// TIA Portal project "DHARMA_1500" (V15)

(* hardware
DEVICE "HMI_DHARMA"  TP1200 Comfort
   slot 0: "KraussMaffeiHMI"  TP1200 Comfort  6AV2 124-0MC01-0AX0  14.0.1.0
   slot 1: "HMI_RT_1"  TP1200 Comfort  6AV2 124-0MC01-0AX0  14.0.1.0
   slot 5: "KraussMaffeiHMI.IE_CP_1"  PROFINET Interface  14.0.1.0
      slot 1: "PROFINET Interface_1"  PROFINET Interface
         slot 1: "Port_1"  Port
         slot 2: "Port_2"  Port
   slot 7: "KraussMaffeiHMI.MPI/DP_CP_1"  MPI/DP Interface  14.0.1.0
DEVICE "S71500/ET200MP station_1"  S7-1500 station
   slot 0: "Rail_0"  Rack  6ES7 590-1***0-0AA0
   slot 1: "PLC_DHARMA"  CPU 1515-2 PN  6ES7 515-2AM01-0AB0  V2.5
      slot 3: "CPU display_1"  6ES7591-1BA00-0AA0
*)

// ===== PLC "PLC_DHARMA"  CPU 1515-2 PN =====

VAR_GLOBAL   // PLC tag table "Standard-Variablentabelle"
   "Sensor_CupIsAtTestshotposition" AT %I18.7 : Bool;   // The cup is at the testhotposition
   "PAW_800_tool_1" AT %QW800 : Word;
   "Tag_3" AT %Q13.2 : Bool;
   "Tag_4" AT %Q13.3 : Bool;
   "Duese_K2_MH01" AT %Q51.2 : Bool;
   "HF_pulse_alarm_GWK1" AT %M1002.4 : Bool;
   "FP_temperingunit_off" AT %M1002.5 : Bool;
   "FP_temperingunit_on" AT %M1002.6 : Bool;
   "With_MC03" AT %M710.0 : Bool;
   "With_MC04" AT %M710.1 : Bool;
   "HF_pulse_alarm_GWK2" AT %M1002.7 : Bool;
   "HF_new_setvalue_Of_ShotData" AT %M701.2 : Bool;
   "HM_Shotend" AT %M50.0 : Bool;
   "TIM_FRA_WDG3" AT %T15 : Timer;
   "TIM_FRA_WDG4" AT %T16 : Timer;
   "T_CupIsAtTestshotposition" AT %T192 : Timer;
END_VAR

VAR_GLOBAL CONSTANT   // PLC tag table "Standard-Variablentabelle"
   "AmountPartShots" : Int := 8;   // Array lenght for UDT 925
   "AmountToolsDB" : Int := 100;   // Array lenght for each DB
   "AmountAllocationAutomatic" : Int := 210;   // Array lenght for DB931 (always 30 Steps)
   "AmountTools" : Int := 200;   // Array lenght for DB930
END_VAR

VAR_GLOBAL   // PLC tag table "E/A- Belegung INput"
   "F_Klima" AT %I4.7 : Bool;   // Malfunction air-condition
   "P_Vacuum_C1" AT %I117.0 : Bool;   // Vacuum reached componet 1
   "P_Vacuum_C2" AT %I117.1 : Bool;   // Vacuum reached componet 2
   "S_BarrelDetection_C1" AT %I111.0 : Bool;   // Special: Barrel exist for the component 1
   "S_BarrelDetection_C2" AT %I112.0 : Bool;   // Special: Barrel exist for the component 2
   "F_Fan_Pump_C1" AT %I110.0 : Bool;   // Fault fuse fan pump component 1
   "F_Fan_Pump_C2" AT %I110.1 : Bool;   // Fault fuse fan pump component 2
   "F_FCFeedingP_C1" AT %I110.4 : Bool;   // Fault frequency drive feed pump component 1
   "F_FCFeedingP_C2" AT %I110.5 : Bool;   // Fault frequency drive feed pump component 2
   "T_Start_Test_C1" AT %I26.3 : Bool;   // Start button for test component 1
   "T_Start_Test_C2" AT %I27.3 : Bool;   // Start button for test component 1
   "T_Stop_Test" AT %I27.2 : Bool;   // Stop button for test component
   "S_OM_Test" AT %I26.2 : Bool;   // Switch for selection operation mode test
   "P_2_MK_Hydr" AT %I2.5 : Bool;   // hydraulic pressure 2 reached
   "ES_GBE_C1" AT %I1.7 : Bool;   // Emergency stop from nucleation component 1
   "F_GBE_C1" AT %I0.5 : Bool;   // Fault Supply nucleation component 1
   "F_GBE_Faulty_C1" AT %I0.6 : Bool;   // Fault Message from nuvleation component 1
   "F_GBE_Ready_C1" AT %I1.3 : Bool;   // Nucleation ready component 1
   "F_FeedPump_C2" AT %I8.6 : Bool;   // Fault filling pump daytank component 2
   "S_DryRun_Feed_C1" AT %I119.2 : Bool;   // Dry run protection feeding pump tank component 1
   "S_DryRun_Feed_C2" AT %I118.3 : Bool;   // Dry run protection feeding pump tank component 2
   "Container_FaultSupply" AT %I10.7 : Bool;   // Faulty power supply containerstaion
   "ES_Door_Robot_01" AT %I13.2 : Bool;   // Emergency stop door robot 1
   "ES_Door_TestShot_01" AT %I18.4 : Bool;   // Emergency stop door testshot robot 1
   "ES_Container_C1" AT %I10.5 : Bool;   // Emergency stop from containerstaion component 1
   "TestShot_MouldExist" AT %I14.4 : Bool;   // Testshot: Mould existing
   "TestShot_Level" AT %I14.5 : Bool;   // Testshot: Filling level
   "S_SelectDoor_Robot_01" AT %I13.0 : Bool;   // Select open door robot 1
   "AS_Door_Robot_01" AT %I13.3 : Bool;   // Automatic stop door robot 1
   "S_QuittDoor_Robot_01" AT %I13.1 : Bool;   // Quitt automatic stop door robot 1
   "S_SelectDoor_TestShot_01" AT %I18.0 : Bool;   // Select open door test shot 1
   "AS_Door_TestShot_01" AT %I18.3 : Bool;   // Automatic stop door test shot 1
   "S_QuittDoor_TestShot_01" AT %I18.1 : Bool;   // Quitt automatic stop door test shot 1
   "AS_RobotInArea1" AT %I12.0 : Bool;   // Save Move (EPS) area 1
   "AS_RobotInArea2" AT %I12.1 : Bool;   // Save Move (EPS) area 2
   "AS_Dryside" AT %I8.7 : Bool;   // Automatic stop from mould carrier 01
   "AS" AT %I12.7 : Bool;   // Emergency stop from dryside
   "F_CoolingDevice" AT %I0.4 : Bool;   // Faulty supply chiller
   "Container_Ready_C1" AT %I10.1 : Bool;   // Signal container is ready for filling daytank component 1
   "Container_Ready_C2" AT %I10.2 : Bool;   // Signal container is ready for filling daytank component 2
   "Container_Fillpump_run_C1" AT %I10.3 : Bool;   // Signal container filling pump is running component 1
   "Container_Fillpump_run_C2" AT %I10.4 : Bool;   // Signal container filling pump is running component 2
   "Container_Faulty" AT %I10.6 : Bool;   // Signal container fault existing
   "F_TraceHeatingM1_C3" AT %I17.3 : Bool;
   "F_FeedingP_C1" AT %I24.0 : Bool;   // Fault Feeding pump component 1
   "F_FeedingP_C2" AT %I25.0 : Bool;   // Fault Feeding pump component 2
   "F_SupplyHeatingM1" AT %I16.0 : Bool;   // Stoerung versorgung heizung
   "F_TraceHeatingM1_C1" AT %I16.1 : Bool;   // Stoerung begleitheizung vorlauf ruecklauf poly
   "F_TraceHeatingM1_C2" AT %I16.2 : Bool;   // Stoerung begleitheizung vorlauf ruecklauf iso
   "F_TraceHeatingM1_C1_2" AT %I16.3 : Bool;
   "F_TraceHeatingM1_C2_2" AT %I16.4 : Bool;
   "F_Robot_01" AT %I12.6 : Bool;   // Fault fuse robot 01
   "F_Airdryer" AT %I0.1 : Bool;   // Fault Airdryer
   "ES_Extern(SGM_or_MC)" AT %I0.0 : Bool;   // Emergency stop from extern (SGM or Mould carrier)
   "F_Fuse_Machine" AT %I0.2 : Bool;   // Fault circuit breakes machine component 1/2
   "F_Fuse_MH" AT %I0.3 : Bool;   // Fault fuse mixinghead
   "ES_Operatingpanel" AT %I1.5 : Bool;   // Emergency stop control panel PUC 08
   "ES_Machine" AT %I1.4 : Bool;   // Emergency stop machine component 1/2
   "Controlvoltage" AT %I0.7 : Bool;   // Control voltage on
   "ES_Robot_01" AT %I12.5 : Bool;   // Emergency stop from robot 01
   "ES_Central" AT %I1.6 : Bool;   // Emergency stop from central
   "S_OM_Manual" AT %I1.0 : Bool;   // Operating mode manual
   "S_OM_Auto" AT %I1.1 : Bool;   // Operating mode automatic
   "T_QuitFault" AT %I1.2 : Bool;
   "F_MK_Hydr" AT %I2.0 : Bool;   // malfunction hydraulicmotor
   "F_Fil_MK_Hydr_VL" AT %I2.1 : Bool;   // hydraulic filter polluted forwardslauf
   "L_Min_Oel_MK_Hydr" AT %I2.2 : Bool;   // hydraulic fill level OK
   "C_Max_Oel_MK_Hydr" AT %I2.3 : Bool;   // Max temperature hydraulic
   "P_MK_Hydr" AT %I2.4 : Bool;   // hydraulic pressure reached
   "C_Cooling_Hydr" AT %I2.6 : Bool;   // Start cooling hydraulic
   "F_Heating" AT %I2.7 : Bool;   // Fault Heating Day tank
   "Select_door_TT" AT %I120.5 : Bool;
   "AS_door_TT" AT %I120.3 : Bool;
   "Quit_door_TT" AT %I120.4 : Bool;
   "F_fuse_vacuum_pump_Seg_1" AT %I121.4 : Bool;
   "F_fuse_vacuum_pump_Seg_2" AT %I122.4 : Bool;
   "F_fuse_vacuum_pump_Seg_3" AT %I123.4 : Bool;
   "F_fuse_vacuum_pump_Seg_4" AT %I124.4 : Bool;
   "Safety_switch_MC_1" AT %I121.2 : Bool;
   "Safety_switch_MC_2" AT %I122.2 : Bool;
   "Safety_switch_MC_3" AT %I123.2 : Bool;
   "Safety_switch_MC_4" AT %I124.2 : Bool;
   "S_Start_TestShot_01" AT %I18.2 : Bool;   // Start automatic test shot 1
   "AS_RobotInArea3" AT %I12.2 : Bool;   // Save Move (EPS) area 3
   "AS_RobotInArea4" AT %I12.3 : Bool;   // Save Move (EPS) area 4
   "AS_RobotInArea5" AT %I18.5 : Bool;   // Save Move (EPS) area 5
   "AS_RobotInArea6" AT %I18.6 : Bool;   // Save Move (EPS) area 6
   "AS_Lightbarrier_back_MC01" AT %I30.3 : Bool;   // Automatic stop light barrier behind MC 1
   "ES_MC02" AT %I30.4 : Bool;   // Emergency stop from mould carrier 2
   "AS_tool_exists_MC02" AT %I30.5 : Bool;   // Automatic stop tool exists mould carrier 2
   "AS_MC02" AT %I30.6 : Bool;   // Automatic stop from mould carrier 2
   "AS_Lightbarrier_back_MC02" AT %I30.7 : Bool;   // Automatic stop light barrier behind MC 2
   "ES_MC03" AT %I31.0 : Bool;   // Emergency stop from mould carrier 3
   "AS_tool_exists_MC03" AT %I31.1 : Bool;   // Automatic stop tool exists mould carrier 3
   "AS_MC03" AT %I31.2 : Bool;   // Automatic stop from mould carrier 3
   "AS_Lightbarrier_back_MC03" AT %I31.3 : Bool;   // Automatic stop light barrier behind MC 3
   "ES_MC04" AT %I31.4 : Bool;   // Emergency stop from mould carrier 4
   "AS_tool_exists_MC04" AT %I31.5 : Bool;   // Automatic stop tool exists mould carrier 4
   "AS_MC04" AT %I31.6 : Bool;   // Automatic stop from mould carrier 4
   "AS_Lightbarrier_back_MC04" AT %I31.7 : Bool;   // Automatic stop light barrier behind MC 4
   "ES_MC01" AT %I30.0 : Bool;   // Emergency stop from mould carrier 1
   "AS_tool_exists_MC01" AT %I30.1 : Bool;   // Automatic stop tool exists mould carrier 1
   "AS_MC01" AT %I30.2 : Bool;   // Automatic stop from mould carrier 1
   "P_air" AT %I19.7 : Bool;   // Pressure air inlet
   "C_Start_Refill_POLY_ON" AT %Q11.1 : Bool;
   "C_Start_Refill_ISO_ON" AT %Q11.2 : Bool;
   "Release_door_TT" AT %Q120.1 : Bool;
   "Selected_door_TT" AT %Q120.0 : Bool;
   "O_vacuum_pump_Seg_1" AT %Q121.1 : Bool;
   "O_vacuum_pump_Seg_2" AT %Q121.2 : Bool;
   "O_vacuum_pump_Seg_3" AT %Q121.3 : Bool;
   "O_vacuum_pump_Seg_4" AT %Q121.4 : Bool;
   "FHM_Takt_Verz_RT1" AT %M900.0 : Bool;
   "HM_FP_Takt_Verz_RT1" AT %M900.1 : Bool;
END_VAR

VAR_GLOBAL   // PLC tag table "E/A- Belegung OUTput"
   "K_ControllVoltageOff" AT %Q0.4 : Bool;
   "K_Stoerung_FT" AT %Q3.0 : Bool;   // malfunction to mouldcarrier
   "K_Schussende_FT" AT %Q3.1 : Bool;   // Shotend an mouldcarrier
   "H_CP_Back_MH1" AT %Q3.2 : Bool;   // MH01: indicator cleaning piston back
   "H_Rel_Foaming_MH1" AT %Q3.3 : Bool;   // MH01: indicator release foaming
   "H_HighPressure_MH1" AT %Q3.4 : Bool;   // MH01: indicator high pressure circulation
   "V_MH_open_MH1" AT %Q115.0 : Bool;   // MH00: Valve mixinghead open
   "V_CP_Forward_MH1" AT %Q115.1 : Bool;   // MH00: valve cleaning piston forward
   "V_PumpVacuum_C1" AT %Q117.0 : Bool;
   "V_PressureVacuum_C1" AT %Q117.1 : Bool;
   "V_PumpVacuum_C2" AT %Q117.2 : Bool;
   "V_PressureVacuum_C2" AT %Q117.3 : Bool;
   "M_CirculationPump_C3" AT %Q118.0 : Bool;   // Circulation Pump net component 3
   "V_PumpVacuum_C3" AT %Q117.4 : Bool;
   "V_PressureVacuum_C3" AT %Q117.5 : Bool;
   "V_PressureVacuum_C4" AT %Q117.7 : Bool;
   "V_Inert_MH1" AT %Q122.6 : Bool;   // MH01: Valve Nitrogen for Inerting
   "V_Inert_Piston_MH1" AT %Q131.5 : Bool;   // MH01: Valve Nitrogen Piston
   "M_Fan_Pump_Net_C1" AT %Q110.0 : Bool;   // Fan pump net component 1
   "M_Fan_Pump_Net_C2" AT %Q110.1 : Bool;   // Fan pump net component 2
   "M_FeedingP_Start_C1" AT %Q24.1 : Bool;   // Feedingpump release frequency drive component 1
   "M_FeedingP_Start_C2" AT %Q25.1 : Bool;   // Feedingpump release frequency drive component 2
   "V_Test_C1" AT %Q26.2 : Bool;   // Valve for test component 1
   "V_Test_C2" AT %Q27.2 : Bool;   // Valve for test component 2
   "H_Test_C1" AT %Q26.3 : Bool;   // Visual information for test component 1
   "H_Test_C2" AT %Q27.3 : Bool;   // Visual information for test component 2
   "V_Pump_2Point_C1" AT %Q5.0 : Bool;   // 2 Point adjustment component pump component 1
   "M_FeedPump_C1" AT %Q27.0 : Bool;   // Valve for feedpump Daytank Component 1
   "M_FeedPump_C2" AT %Q26.0 : Bool;   // Valve for feedpump Daytank Component 2
   "V_Pump_2Point_C2" AT %Q5.1 : Bool;   // 2 Point adjustment component pump component 2
   "V_OpenDoor_Robot_01" AT %Q13.1 : Bool;   // Clamping valve door robot 01
   "H_ReleaseDoor_Robot_01" AT %Q13.0 : Bool;   // Light door robot 01
   "V_OpenDoor_TestShot_01" AT %Q18.0 : Bool;   // Clamping valve door test shot 01
   "H_AutoStopQuit" AT %Q0.3 : Bool;   // Indicator auto stop acknowledged
   "H_ReleaseDoor_TestShot_01" AT %Q18.1 : Bool;   // Light door test shot 01
   "V_P_builtup_MH_Hydr_M1" AT %Q1.1 : Bool;   // Hydraulic pressur built up mixinhead 1
   "V_Cooling_Hydr" AT %Q1.2 : Bool;   // Hydraulic 1 valve for oil cooling
   "M_MH_Hydr_Net_M1" AT %Q1.0 : Bool;   // Hydraulic motor net mixinghead 1
   "H_Fault_lamp_M1" AT %Q0.0 : Bool;   // Visual fault warning M1
   "H_Fault_horn_M1" AT %Q0.1 : Bool;   // Acustical fault warning M1
   "H_Ready_for_Operation" AT %Q0.2 : Bool;
   "H_TestShot_active_01" AT %Q18.2 : Bool;   // Automatic test shot is running 01
END_VAR

VAR_GLOBAL   // PLC tag table "I/O- Pentan"
   "E_Voralarm_Pentan" AT %I116.0 : Bool;   // Pentan: Pre alarm (20%) pentan
   "P_Voralarm_Stickstoff" AT %I116.1 : Bool;   // Pentan: Pre alarm nitrogen
   "P_Alarm_Stickstoff" AT %I116.2 : Bool;   // Pentan: Alarm nitrogen
   "P_Alarm_VersorgungN" AT %I116.3 : Bool;   // Pentan: Alarm nitrogen supply
   "E_Absaugung_bereit" AT %I116.4 : Bool;   // Pentan: Exhaust system ready
   "E_Pentanpumpe_laeuft" AT %I116.5 : Bool;   // Pentan: Pump pentan running
   "E_Pentamix_Ready" AT %I116.6 : Bool;   // Pentan: Pentamix ready for supply
   "ES_Pentamix" AT %I116.7 : Bool;
   "P_Nitrogen_Inerting_OK" AT %I17.6 : Bool;   // Nitrogen pressure for Inerting ok
   "Flow_Nitrogen Inert_OK" AT %I17.7 : Bool;   // Nitrogen flow after start inerting ok
   "K_Machine_Running" AT %Q116.0 : Bool;   // Pentan: Signal machine running to gas warning desk
   "K_Request_WeekendMode" AT %Q116.1 : Bool;   // Pentan: Request for weekend mode to gas warning desk
   "V_Fass_Pentan1" AT %Q1101.6 : Bool;
   "V_ChargingTank_C1_2" AT %Q22.4 : Bool;   // Filling valve 2 tank component 1
END_VAR

VAR_GLOBAL   // PLC tag table "I/O- PN Modul Flow Output"
   "V_ChargingTank_C2_2" AT %Q22.3 : Bool;   // Filling valve 2 tank component 1
   "M_Pump_Net_C1" AT %Q20.0 : Bool;   // Pump net componet 1
   "M_Pump_Start_C1" AT %Q20.1 : Bool;   // Pump release frequency drive component 1
   "M_Platefilter_C1" AT %Q20.7 : Bool;   // Platefilter net componet 1
   "M_Pump_Net_C2" AT %Q22.0 : Bool;   // Pump net component 2
   "M_Pump_Start_C2" AT %Q22.1 : Bool;   // Pump release frequency drive component 2
   "M_Platefilter_C2" AT %Q22.7 : Bool;   // Platefilter net component 2
   "V_HP_Heater_Cooling_C1" AT %Q21.6 : Bool;   // Valve for cooling high pressure heatexchanger component 1
   "V_HP_Heater_Bypass_C1" AT %Q80.6 : Bool;   // Valve for bypass high pressure heatexchanger component 1
   "V_HP_Heater_Cooling_C2" AT %Q23.6 : Bool;   // Valve for cooling high pressure heatexchanger component 2
   "K_Filling_Tank_C2_TL" AT %Q23.7 : Bool;   // Potential-free contact for filling Tank component 2 from another source
   "M_FU_Start_RW_K1" AT %Q21.1 : Bool;   // Agitator release frequency drive component 1
   "M_FU_Start_RW_K2" AT %Q23.1 : Bool;   // Agitator release frequency drive component 2
   "M_FeedingP_C1" AT %Q24.0 : Bool;   // Feeding pump net component 2
   "M_FeedingP_C2" AT %Q25.0 : Bool;   // Feeding pump net component 2
   "K_Filling_Tank_C2" AT %Q23.3 : Bool;   // Potential-free contact for filling Tank component 2
   "K_Filling_Tank_C1" AT %Q21.3 : Bool;   // Potential-free contact for filling Tank component 1
   "M_AgitatorBarrel_C1" AT %Q20.4 : Bool;   // Agitator barrel net component 1
   "M_Agitator_C1" AT %Q21.0 : Bool;   // Agitator net component 1
   "K_HeatingTank_C1" AT %Q20.2 : Bool;   // Heating Day tank net componet 1
   "V_Coolingwater_C1" AT %Q21.4 : Bool;   // Valve cooling water tank component 1
   "V_ChargingTank_C1" AT %Q21.2 : Bool;   // Filling valve tank component 1
   "V_Barrel_C1" AT %Q20.5 : Bool;   // Valve barrel station component 1
   "V_Heatexchanger_C1" AT %Q21.5 : Bool;   // heat exchangerValve Poly
   "V_Barrel_C2" AT %Q22.5 : Bool;   // Valve barrel station component 2
   "V_Heatexchanger_C2" AT %Q23.5 : Bool;   // heat exchangerValve component 2
   "V_Coolingwater_C2" AT %Q23.4 : Bool;   // Valve cooling water component 2
   "K_HeatingTank_C2" AT %Q22.2 : Bool;   // Heating Day tank net componet 2
   "V_ChargingTank_C2" AT %Q23.2 : Bool;   // Filling valve component 2
   "M_Agitator_C2" AT %Q23.0 : Bool;   // Agitator net component 2
   "V_LowPressure_Circ_C1" AT %Q20.6 : Bool;   // Low pressure circulation component 1
   "V_LowPressure_Circ_C2" AT %Q22.6 : Bool;   // Low pressure circulation component 2
END_VAR

VAR_GLOBAL   // PLC tag table "I/O- PN Modul Flow Input"
   "F_FC_Pump_C1" AT %I20.2 : Bool;   // Fault frequency drive componet 1
   "F_Pump_C1" AT %I20.3 : Bool;   // Fault pump componet 1
   "P_Prepressure_Pump_C1" AT %I20.4 : Bool;   // Pre pressure pump componet 1
   "P_Min_C1" AT %I20.5 : Bool;   // Min. pressure pump componet 1
   "P_Max_C1" AT %I20.6 : Bool;   // Max. pressure pump componet 1
   "F_Platefilter_C1" AT %I20.7 : Bool;   // Fault Platefilter component 1
   "F_FC_Agitator_C1" AT %I21.1 : Bool;   // Malfunction frequency converter agitator component 1
   "F_FC_Pump_C2" AT %I22.2 : Bool;   // Fault frequency drive componet 2
   "F_Pump_C2" AT %I22.3 : Bool;   // Fault pump componet 2
   "P_Prepressure_Pump_C2" AT %I22.4 : Bool;   // Pre pressure pump componet 2
   "P_Min_C2" AT %I22.5 : Bool;   // Min. pressure pump componet 2
   "F_Platefilter_C2" AT %I22.7 : Bool;   // Fault Platefilter component 2
   "P_Max_C2" AT %I22.6 : Bool;   // Max. pressure pump componet 2
   "F_FC_Agitator_C2" AT %I23.1 : Bool;   // Malfunction frequency converter agitator component 2
   "F_Agitator_C1" AT %I21.0 : Bool;   // Fault agitator componet 1
   "F_Temperiergeraet_C1" AT %I21.7 : Bool;   // Malfunction temperature stabilizer component 1
   "L_Tank_min_C1" AT %I21.2 : Bool;   // Min fill level tank componet 1
   "L_Tank_start_C1" AT %I21.3 : Bool;   // Start refilling level tank componet 1
   "L_Tank_stop_C1" AT %I21.4 : Bool;   // Stop refilling level tank componet 1
   "L_DT_max_C1" AT %I21.5 : Bool;   // Max. Filling level componet 1
   "L_DripTray_C1" AT %I21.6 : Bool;   // Max. level drip tray componet 1
   "F_Agitator_C2" AT %I23.0 : Bool;   // Fault agitator componet 2
   "F_Temperiergeraet_C2" AT %I23.7 : Bool;   // Malfunction temperature stabilizer component 2
   "L_Tank_min_C2" AT %I23.2 : Bool;   // Min fill level componet 2
   "L_Tank_start_C2" AT %I23.3 : Bool;   // Start refilling level componet 2
   "L_Tank_stop_C2" AT %I23.4 : Bool;   // Stop refilling level componet 2
   "L_DT_max_C2" AT %I23.5 : Bool;   // Max. Filling level componet 2
   "L_DripTray_C2" AT %I23.6 : Bool;   // Max. level drip tray componet 2
   "Kracht_C1_A_Flowrate" AT %I20.0 : Bool;
   "Kracht_C1_B_Flowrate" AT %I20.1 : Bool;
   "Kracht_C2_A_Flowrate" AT %I22.0 : Bool;
   "Kracht_C2_B_Flowrate" AT %I22.1 : Bool;
END_VAR

VAR_GLOBAL   // PLC tag table "I/O- PN Modul Mixinghead Output"
   "V_SWU_MH01" AT %Q50.5 : Bool;   // MH01: Valve switch over unit
   "H_Shotcounter_MH01" AT %Q52.7 : Bool;   // MH01: shot counter
   "V_CP_Forward_MH01" AT %Q50.4 : Bool;   // MH01: valve cleaning piston forward
   "H_CP_Back_MH01" AT %Q52.4 : Bool;   // MH01: indicator cleaning piston back
   "H_Rel_Foaming_MH01" AT %Q52.6 : Bool;   // MH01: indicator release foaming
   "H_HighPressure_MH01" AT %Q52.5 : Bool;   // MH01: indicator high pressure circulation
   "K_Fault_MC01" AT %Q50.6 : Bool;   // MH01: malfunction PU-machine to mouldcarrier
   "K_ShotEnd_MC01" AT %Q50.7 : Bool;   // MH01: Shotend PU-machine to mouldcarrier
   "V_MH_open_MH01" AT %Q50.0 : Bool;   // MH01: Valve mixinghead open
   "V_LowPressure_Circ_MH01" AT %Q53.7 : Bool;   // MH01: low pressure circulation Poly/ Iso
   "V_MH_open_MH02" AT %Q54.0 : Bool;   // MH01: Valve mixinghead open
   "V_CP_Forward_MH02" AT %Q54.4 : Bool;   // MH01: valve cleaning piston forward
   "V_SWU_MH02" AT %Q54.5 : Bool;   // MH01: Valve switch over unit
   "K_Fault_MC02" AT %Q54.6 : Bool;   // MH01: malfunction PU-machine to mouldcarrier
   "K_ShotEnd_MC02" AT %Q54.7 : Bool;   // MH01: Shotend PU-machine to mouldcarrier
   "H_CP_Back_MH02" AT %Q56.4 : Bool;   // MH01: indicator cleaning piston back
   "H_HighPressure_MH02" AT %Q56.5 : Bool;   // MH01: indicator high pressure circulation
   "H_Rel_Foaming_MH02" AT %Q56.6 : Bool;   // MH01: indicator release foaming
   "H_Shotcounter_MH02" AT %Q56.7 : Bool;   // MH01: shot counter
   "V_LowPressure_Circ_MH02" AT %Q57.7 : Bool;   // MH01: low pressure circulation Poly/ Iso
   "V_MH_open_MH03" AT %Q58.0 : Bool;   // MH01: Valve mixinghead open
   "V_CP_Forward_MH03" AT %Q58.4 : Bool;   // MH01: valve cleaning piston forward
   "V_SWU_MH03" AT %Q58.5 : Bool;   // MH01: Valve switch over unit
   "K_Fault_MC03" AT %Q58.6 : Bool;   // MH01: malfunction PU-machine to mouldcarrier
   "K_ShotEnd_MC03" AT %Q58.7 : Bool;   // MH01: Shotend PU-machine to mouldcarrier
   "H_CP_Back_MH03" AT %Q60.4 : Bool;   // MH01: indicator cleaning piston back
   "H_HighPressure_MH03" AT %Q60.5 : Bool;   // MH01: indicator high pressure circulation
   "H_Rel_Foaming_MH03" AT %Q60.6 : Bool;   // MH01: indicator release foaming
   "H_Shotcounter_MH03" AT %Q60.7 : Bool;   // MH01: shot counter
   "V_LowPressure_Circ_MH03" AT %Q61.7 : Bool;   // MH01: low pressure circulation Poly/ Iso
   "V_MH_open_MH04" AT %Q62.0 : Bool;   // MH01: Valve mixinghead open
   "V_CP_Forward_MH04" AT %Q62.4 : Bool;   // MH01: valve cleaning piston forward
   "V_SWU_MH04" AT %Q62.5 : Bool;   // MH01: Valve switch over unit
   "K_Fault_MC04" AT %Q62.6 : Bool;   // MH01: malfunction PU-machine to mouldcarrier
   "K_ShotEnd_MC04" AT %Q62.7 : Bool;   // MH01: Shotend PU-machine to mouldcarrier
   "H_CP_Back_MH04" AT %Q64.4 : Bool;   // MH01: indicator cleaning piston back
   "H_HighPressure_MH04" AT %Q64.5 : Bool;   // MH01: indicator high pressure circulation
   "H_Rel_Foaming_MH04" AT %Q64.6 : Bool;   // MH01: indicator release foaming
   "H_Shotcounter_MH04" AT %Q64.7 : Bool;   // MH01: shot counter
   "V_LowPressure_Circ_MH04" AT %Q65.7 : Bool;   // MH01: low pressure circulation Poly/ Iso
   "V_MH_open_MH05" AT %Q66.0 : Bool;   // MH01: Valve mixinghead open
   "V_CP_Forward_MH05" AT %Q66.4 : Bool;   // MH01: valve cleaning piston forward
   "V_SWU_MH05" AT %Q66.5 : Bool;   // MH01: Valve switch over unit
   "K_Fault_MC05" AT %Q66.6 : Bool;   // MH01: malfunction PU-machine to mouldcarrier
   "K_ShotEnd_MC05" AT %Q66.7 : Bool;   // MH01: Shotend PU-machine to mouldcarrier
   "H_CP_Back_MH05" AT %Q68.4 : Bool;   // MH01: indicator cleaning piston back
   "H_HighPressure_MH05" AT %Q68.5 : Bool;   // MH01: indicator high pressure circulation
   "H_Rel_Foaming_MH05" AT %Q68.6 : Bool;   // MH01: indicator release foaming
   "H_Shotcounter_MH05" AT %Q68.7 : Bool;   // MH01: shot counter
   "V_LowPressure_Circ_MH05" AT %Q69.7 : Bool;   // MH01: low pressure circulation Poly/ Iso
   "V_MH_open_MH06" AT %Q70.0 : Bool;   // MH01: Valve mixinghead open
   "V_CP_Forward_MH06" AT %Q70.4 : Bool;   // MH01: valve cleaning piston forward
   "V_SWU_MH06" AT %Q70.5 : Bool;   // MH01: Valve switch over unit
   "K_Fault_MC06" AT %Q70.6 : Bool;   // MH01: malfunction PU-machine to mouldcarrier
   "K_ShotEnd_MC06" AT %Q70.7 : Bool;   // MH01: Shotend PU-machine to mouldcarrier
   "H_CP_Back_MH06" AT %Q72.4 : Bool;   // MH01: indicator cleaning piston back
   "H_HighPressure_MH06" AT %Q72.5 : Bool;   // MH01: indicator high pressure circulation
   "H_Rel_Foaming_MH06" AT %Q72.6 : Bool;   // MH01: indicator release foaming
   "H_Shotcounter_MH06" AT %Q72.7 : Bool;   // MH01: shot counter
   "V_LowPressure_Circ_MH06" AT %Q73.7 : Bool;   // MH01: low pressure circulation Poly/ Iso
   "V_MH_open_MH07" AT %Q74.0 : Bool;   // MH01: Valve mixinghead open
   "V_CP_Forward_MH07" AT %Q74.4 : Bool;   // MH01: valve cleaning piston forward
   "V_SWU_MH07" AT %Q74.5 : Bool;   // MH01: Valve switch over unit
   "K_Fault_MC07" AT %Q74.6 : Bool;   // MH01: malfunction PU-machine to mouldcarrier
   "K_ShotEnd_MC07" AT %Q74.7 : Bool;   // MH01: Shotend PU-machine to mouldcarrier
   "H_CP_Back_MH07" AT %Q76.4 : Bool;   // MH01: indicator cleaning piston back
   "H_HighPressure_MH07" AT %Q76.5 : Bool;   // MH01: indicator high pressure circulation
   "H_Rel_Foaming_MH07" AT %Q76.6 : Bool;   // MH01: indicator release foaming
   "H_Shotcounter_MH07" AT %Q76.7 : Bool;   // MH01: shot counter
   "V_LowPressure_Circ_MH07" AT %Q77.7 : Bool;   // MH01: low pressure circulation Poly/ Iso
   "V_MH_open_MH08" AT %Q78.0 : Bool;   // MH01: Valve mixinghead open
   "V_CP_Forward_MH08" AT %Q78.4 : Bool;   // MH01: valve cleaning piston forward
   "V_SWU_MH08" AT %Q78.5 : Bool;   // MH01: Valve switch over unit
   "K_Fault_MC08" AT %Q78.6 : Bool;   // MH01: malfunction PU-machine to mouldcarrier
   "K_ShotEnd_MC08" AT %Q78.7 : Bool;   // MH01: Shotend PU-machine to mouldcarrier
   "H_CP_Back_MH08" AT %Q80.4 : Bool;   // MH01: indicator cleaning piston back
   "H_HighPressure_MH08" AT %Q80.5 : Bool;   // MH01: indicator high pressure circulation
   "K_Filling_Tank_C1_TL" AT %Q21.7 : Bool;   // Potential-free contact for filling Tank component 1 from another source
   "H_Shotcounter_MH08" AT %Q80.7 : Bool;   // MH01: shot counter
   "V_LowPressure_Circ_MH08" AT %Q81.7 : Bool;   // MH01: low pressure circulation Poly/ Iso
   "V_MH_open_MH09" AT %Q82.0 : Bool;   // MH01: Valve mixinghead open
   "V_CP_Forward_MH09" AT %Q82.4 : Bool;   // MH01: valve cleaning piston forward
   "V_SWU_MH09" AT %Q82.5 : Bool;   // MH01: Valve switch over unit
   "K_Fault_MC09" AT %Q82.6 : Bool;   // MH01: malfunction PU-machine to mouldcarrier
   "K_ShotEnd_MC09" AT %Q82.7 : Bool;   // MH01: Shotend PU-machine to mouldcarrier
   "H_CP_Back_MH09" AT %Q84.4 : Bool;   // MH01: indicator cleaning piston back
   "H_HighPressure_MH09" AT %Q84.5 : Bool;   // MH01: indicator high pressure circulation
   "H_Rel_Foaming_MH09" AT %Q84.6 : Bool;   // MH01: indicator release foaming
   "H_Shotcounter_MH09" AT %Q84.7 : Bool;   // MH01: shot counter
   "V_LowPressure_Circ_MH09" AT %Q85.7 : Bool;   // MH01: low pressure circulation Poly/ Iso
   "V_MH_open_MH10" AT %Q86.0 : Bool;   // MH01: Valve mixinghead open
   "V_CP_Forward_MH10" AT %Q86.4 : Bool;   // MH01: valve cleaning piston forward
   "V_SWU_MH10" AT %Q86.5 : Bool;   // MH01: Valve switch over unit
   "K_Fault_MC10" AT %Q86.6 : Bool;   // MH01: malfunction PU-machine to mouldcarrier
   "K_ShotEnd_MC10" AT %Q86.7 : Bool;   // MH01: Shotend PU-machine to mouldcarrier
   "H_CP_Back_MH10" AT %Q88.4 : Bool;   // MH01: indicator cleaning piston back
   "H_HighPressure_MH10" AT %Q88.5 : Bool;   // MH01: indicator high pressure circulation
   "H_Rel_Foaming_MH10" AT %Q88.6 : Bool;   // MH01: indicator release foaming
   "H_Shotcounter_MH10" AT %Q88.7 : Bool;   // MH01: shot counter
   "V_LowPressure_Circ_MH10" AT %Q95.7 : Bool;   // MH01: low pressure circulation Poly/ Iso
   "V_Bypass_C1" AT %Q51.1 : Bool;
   "V_Bypass_C2" AT %Q51.3 : Bool;
   "Duese_K1_MH01" AT %Q51.0 : Bool;
END_VAR

VAR_GLOBAL   // PLC tag table "I/O- PN Modul Mixinghead Input"
   "T_CP_forward_MH01" AT %I52.3 : Bool;   // MH01: Button cleaning piston forwards
   "T_CP_back_MH01" AT %I52.4 : Bool;   // MH01: Button cleaning piston back
   "S_ProgrNo_Bit40_MH01" AT %I51.6 : Bool;   // MH01: preselection program no. *10 MH BIT 2
   "P_Min_Air" AT %I53.6 : Bool;   // MH01: Min. Druck Reinigungsluft
   "P_Max_Air" AT %I53.7 : Bool;   // MH01: Max. Druck Reinigungsluft
   "S_ProgrNo_Bit80_MH01" AT %I51.7 : Bool;   // MH01: preselection program no. *10 MH BIT 3
   "ES_OP_Panel_MH01" AT %I50.2 : Bool;   // MH01: Emergency stop operating panel mixinghead
   "IPS_MH_MH01" AT %I50.0 : Bool;   // MH01: Inductive proximity switch mixinghead
   "IPS_CP_MH01" AT %I50.1 : Bool;   // MH01: Inductive proximity switch cleaning piston mixinghead
   "K_PreparationFoamingMC01" AT %I50.6 : Bool;   // MH01: preparation foaming from mouldcarrier
   "K_FoamingReleaseMC01" AT %I50.7 : Bool;   // MH01: shot release from mouldcarrier
   "S_Rel_SWU_MH01" AT %I52.2 : Bool;   // MH01: release switch over unit
   "S_Manuel_MH01" AT %I52.0 : Bool;   // MH01: operation mode manual
   "S_Automatic_MH01" AT %I52.1 : Bool;   // MH01: operation mode automatic
   "T_Highpressure_MH01" AT %I52.5 : Bool;   // MH01: Button high pressure circulation
   "S_ProgrNo_Bit20_MH01" AT %I51.5 : Bool;   // MH01: preselection program no. *10 MH BIT 1
   "S_ProgrNo_Bit10_MH01" AT %I51.4 : Bool;   // MH01: preselection program no. *10 MH BIT 0
   "S_ProgNoSelectMH01" AT %IB51 : Byte;   // MH01: preselection program no. MH
   "S_ProgrNo_Bit0_MH01" AT %I51.0 : Bool;   // MH01: preselection program no. MH BIT 0
   "S_ProgrNo_Bit1_MH01" AT %I51.1 : Bool;   // MH01: preselection program no. MH BIT 1
   "S_ProgrNo_Bit2_MH01" AT %I51.2 : Bool;   // MH01: preselection program no. MH BIT 2
   "S_ProgrNo_Bit3_MH01" AT %I51.3 : Bool;   // MH01: preselection program no. MH BIT 3
   "T_Start_MH01" AT %I52.6 : Bool;   // MH01: Button Start foaming
   "T_Stop_MH01" AT %I52.7 : Bool;   // MH01: Button Stop foaming
   "T_BreakeOpen_MH01" AT %I53.5 : Bool;   // MH01: Button to open the boom brake
   "IPS_MH_MH02" AT %I54.0 : Bool;   // MH02: Inductive proximity switch mixinghead
   "IPS_CP_MH02" AT %I54.1 : Bool;   // MH02: Inductive proximity switch cleaning piston mixinghead
   "ES_OP_Panel_MH02" AT %I54.2 : Bool;   // MH02: Emergency stop operating panel mixinghead
   "K_PreparationFoamingMC02" AT %I54.6 : Bool;   // MH02: preparation foaming from mouldcarrier
   "K_FoamingReleaseMC02" AT %I54.7 : Bool;   // MH02: shot release from mouldcarrier
   "S_ProgNoSelectMH02" AT %IB55 : Byte;   // MH02: preselection program no. MH
   "S_ProgrNo_Bit0_MH02" AT %I55.0 : Bool;   // MH02: preselection program no. MH BIT 0
   "S_ProgrNo_Bit1_MH02" AT %I55.1 : Bool;   // MH02: preselection program no. MH BIT 1
   "S_ProgrNo_Bit2_MH02" AT %I55.2 : Bool;   // MH02: preselection program no. MH BIT 2
   "S_ProgrNo_Bit3_MH02" AT %I55.3 : Bool;   // MH02: preselection program no. MH BIT 3
   "S_ProgrNo_Bit10_MH02" AT %I55.4 : Bool;   // MH02: preselection program no. *10 MH BIT 0
   "S_ProgrNo_Bit20_MH02" AT %I55.5 : Bool;   // MH02: preselection program no. *10 MH BIT 1
   "S_ProgrNo_Bit40_MH02" AT %I55.6 : Bool;   // MH02: preselection program no. *10 MH BIT 2
   "S_ProgrNo_Bit80_MH02" AT %I55.7 : Bool;   // MH02: preselection program no. *10 MH BIT 3
   "S_Manuel_MH02" AT %I724.0 : Bool;   // MH02: operation mode manual
   "S_Automatic_MH02" AT %I724.1 : Bool;   // MH02: operation mode automatic
   "S_Rel_SWU_MH02" AT %I724.2 : Bool;   // MH02: release switch over unit
   "T_CP_forward_MH02" AT %I724.3 : Bool;   // MH02: Button cleaning piston forwards
   "T_CP_back_MH02" AT %I724.4 : Bool;   // MH02: Button cleaning piston back
   "T_Highpressure_MH02" AT %I724.5 : Bool;   // MH02: Button high pressure circulation
   "T_Start_MH02" AT %I724.6 : Bool;   // MH02: Button Start foaming
   "T_Stop_MH02" AT %I724.7 : Bool;   // MH02: Button Stop foaming
   "P_Min_Air_MH02" AT %I725.6 : Bool;   // MH02: Min. Druck Reinigungsluft
   "P_Max_Air_MH02" AT %I725.7 : Bool;   // MH02: Max. Druck Reinigungsluft
   "T_BreakeOpen_MH02" AT %I725.5 : Bool;   // MH02: Button to open the boom brake
   "IPS_MH_MH03" AT %I726.0 : Bool;   // MH03: Inductive proximity switch mixinghead
   "IPS_CP_MH03" AT %I726.1 : Bool;   // MH03: Inductive proximity switch cleaning piston mixinghead
   "ES_OP_Panel_MH03" AT %I726.2 : Bool;   // MH03: Emergency stop operating panel mixinghead
   "K_PreparationFoamingMC03" AT %I726.6 : Bool;   // MH03: preparation foaming from mouldcarrier
   "K_FoamingReleaseMC03" AT %I726.7 : Bool;   // MH03: shot release from mouldcarrier
   "S_ProgNoSelectMH03" AT %IB727 : Byte;   // MH03: preselection program no. MH
   "S_ProgrNo_Bit0_MH03" AT %I727.0 : Bool;   // MH03: preselection program no. MH BIT 0
   "S_ProgrNo_Bit1_MH03" AT %I727.1 : Bool;   // MH03: preselection program no. MH BIT 1
   "S_ProgrNo_Bit2_MH03" AT %I727.2 : Bool;   // MH03: preselection program no. MH BIT 2
   "S_ProgrNo_Bit3_MH03" AT %I727.3 : Bool;   // MH03: preselection program no. MH BIT 3
   "S_ProgrNo_Bit10_MH03" AT %I727.4 : Bool;   // MH03: preselection program no. *10 MH BIT 0
   "S_ProgrNo_Bit20_MH03" AT %I727.5 : Bool;   // MH03: preselection program no. *10 MH BIT 1
   "S_ProgrNo_Bit40_MH03" AT %I727.6 : Bool;   // MH03: preselection program no. *10 MH BIT 2
   "S_ProgrNo_Bit80_MH03" AT %I727.7 : Bool;   // MH03: preselection program no. *10 MH BIT 3
   "S_Manuel_MH03" AT %I728.0 : Bool;   // MH03: operation mode manual
   "S_Automatic_MH03" AT %I728.1 : Bool;   // MH03: operation mode automatic
   "S_Rel_SWU_MH03" AT %I728.2 : Bool;   // MH03: release switch over unit
   "T_CP_forward_MH03" AT %I728.3 : Bool;   // MH03: Button cleaning piston forwards
   "T_CP_back_MH03" AT %I728.4 : Bool;   // MH03: Button cleaning piston back
   "T_Highpressure_MH03" AT %I728.5 : Bool;   // MH03: Button high pressure circulation
   "T_Start_MH03" AT %I728.6 : Bool;   // MH03: Button Start foaming
   "T_Stop_MH03" AT %I728.7 : Bool;   // MH03: Button Stop foaming
   "P_Min_Air_MH03" AT %I729.6 : Bool;   // MH03: Min. Druck Reinigungsluft
   "P_Max_Air_MH03" AT %I729.7 : Bool;   // MH03: Max. Druck Reinigungsluft
   "T_BreakeOpen_MH03" AT %I729.5 : Bool;   // MH03: Button to open the boom brake
   "IPS_MH_MH04" AT %I730.0 : Bool;   // MH03: Inductive proximity switch mixinghead
   "IPS_CP_MH04" AT %I730.1 : Bool;   // MH03: Inductive proximity switch cleaning piston mixinghead
   "ES_OP_Panel_MH04" AT %I730.2 : Bool;   // MH03: Emergency stop operating panel mixinghead
   "K_PreparationFoamingMC04" AT %I730.6 : Bool;   // MH03: preparation foaming from mouldcarrier
   "K_FoamingReleaseMC04" AT %I730.7 : Bool;   // MH03: shot release from mouldcarrier
   "S_ProgNoSelectMH04" AT %IB731 : Byte;   // MH03: preselection program no. MH
   "S_ProgrNo_Bit0_MH04" AT %I731.0 : Bool;   // MH03: preselection program no. MH BIT 0
   "S_ProgrNo_Bit1_MH04" AT %I731.1 : Bool;   // MH03: preselection program no. MH BIT 1
   "S_ProgrNo_Bit2_MH04" AT %I731.2 : Bool;   // MH03: preselection program no. MH BIT 2
   "S_ProgrNo_Bit3_MH04" AT %I731.3 : Bool;   // MH03: preselection program no. MH BIT 3
   "S_ProgrNo_Bit10_MH04" AT %I731.4 : Bool;   // MH03: preselection program no. *10 MH BIT 0
   "S_ProgrNo_Bit20_MH04" AT %I731.5 : Bool;   // MH03: preselection program no. *10 MH BIT 1
   "S_ProgrNo_Bit40_MH04" AT %I731.6 : Bool;   // MH03: preselection program no. *10 MH BIT 2
   "S_ProgrNo_Bit80_MH04" AT %I731.7 : Bool;   // MH03: preselection program no. *10 MH BIT 3
   "S_Manuel_MH04" AT %I732.0 : Bool;   // MH03: operation mode manual
   "S_Automatic_MH04" AT %I732.1 : Bool;   // MH03: operation mode automatic
   "S_Rel_SWU_MH04" AT %I732.2 : Bool;   // MH03: release switch over unit
   "T_CP_forward_MH04" AT %I732.3 : Bool;   // MH03: Button cleaning piston forwards
   "T_CP_back_MH04" AT %I732.4 : Bool;   // MH03: Button cleaning piston back
   "T_Highpressure_MH04" AT %I732.5 : Bool;   // MH03: Button high pressure circulation
   "T_Start_MH04" AT %I732.6 : Bool;   // MH03: Button Start foaming
   "T_Stop_MH04" AT %I732.7 : Bool;   // MH03: Button Stop foaming
   "P_Min_Air_MH04" AT %I733.6 : Bool;   // MH03: Min. Druck Reinigungsluft
   "P_Max_Air_MH04" AT %I733.7 : Bool;   // MH03: Max. Druck Reinigungsluft
   "T_BreakeOpen_MH04" AT %I733.5 : Bool;   // MH03: Button to open the boom brake
   "IPS_MH_MH05" AT %I66.0 : Bool;   // MH03: Inductive proximity switch mixinghead
   "IPS_CP_MH05" AT %I66.1 : Bool;   // MH03: Inductive proximity switch cleaning piston mixinghead
   "ES_OP_Panel_MH05" AT %I66.2 : Bool;   // MH03: Emergency stop operating panel mixinghead
   "K_PreparationFoamingMC05" AT %I66.6 : Bool;   // MH03: preparation foaming from mouldcarrier
   "K_FoamingReleaseMC05" AT %I66.7 : Bool;   // MH03: shot release from mouldcarrier
   "S_ProgNoSelectMH05" AT %IB67 : Byte;   // MH03: preselection program no. MH
   "S_ProgrNo_Bit0_MH05" AT %I67.0 : Bool;   // MH03: preselection program no. MH BIT 0
   "S_ProgrNo_Bit1_MH05" AT %I67.1 : Bool;   // MH03: preselection program no. MH BIT 1
   "S_ProgrNo_Bit2_MH05" AT %I67.2 : Bool;   // MH03: preselection program no. MH BIT 2
   "S_ProgrNo_Bit3_MH05" AT %I67.3 : Bool;   // MH03: preselection program no. MH BIT 3
   "S_ProgrNo_Bit10_MH05" AT %I67.4 : Bool;   // MH03: preselection program no. *10 MH BIT 0
   "S_ProgrNo_Bit20_MH05" AT %I67.5 : Bool;   // MH03: preselection program no. *10 MH BIT 1
   "S_ProgrNo_Bit40_MH05" AT %I67.6 : Bool;   // MH03: preselection program no. *10 MH BIT 2
   "S_ProgrNo_Bit80_MH05" AT %I67.7 : Bool;   // MH03: preselection program no. *10 MH BIT 3
   "S_Manuel_MH05" AT %I68.0 : Bool;   // MH03: operation mode manual
   "S_Automatic_MH05" AT %I68.1 : Bool;   // MH03: operation mode automatic
   "S_Rel_SWU_MH05" AT %I68.2 : Bool;   // MH03: release switch over unit
   "T_CP_forward_MH05" AT %I68.3 : Bool;   // MH03: Button cleaning piston forwards
   "T_CP_back_MH05" AT %I68.4 : Bool;   // MH03: Button cleaning piston back
   "T_Highpressure_MH05" AT %I68.5 : Bool;   // MH03: Button high pressure circulation
   "T_Start_MH05" AT %I68.6 : Bool;   // MH03: Button Start foaming
   "T_Stop_MH05" AT %I68.7 : Bool;   // MH03: Button Stop foaming
   "P_Min_Air_MH05" AT %I69.6 : Bool;   // MH03: Min. Druck Reinigungsluft
   "P_Max_Air_MH05" AT %I69.7 : Bool;   // MH03: Max. Druck Reinigungsluft
   "T_BreakeOpen_MH05" AT %I69.5 : Bool;   // MH03: Button to open the boom brake
   "IPS_MH_MH06" AT %I70.0 : Bool;   // MH06: Inductive proximity switch mixinghead
   "IPS_CP_MH06" AT %I70.1 : Bool;   // MH06: Inductive proximity switch cleaning piston mixinghead
   "ES_OP_Panel_MH06" AT %I70.2 : Bool;   // MH06: Emergency stop operating panel mixinghead
   "K_PreparationFoamingMC06" AT %I70.6 : Bool;   // MH06: preparation foaming from mouldcarrier
   "K_FoamingReleaseMC06" AT %I70.7 : Bool;   // MH06: shot release from mouldcarrier
   "S_ProgNoSelectMH06" AT %IB71 : Byte;   // MH06: preselection program no. MH
   "S_ProgrNo_Bit0_MH06" AT %I71.0 : Bool;   // MH06: preselection program no. MH BIT 0
   "S_ProgrNo_Bit1_MH06" AT %I71.1 : Bool;   // MH06: preselection program no. MH BIT 1
   "S_ProgrNo_Bit2_MH06" AT %I71.2 : Bool;   // MH06: preselection program no. MH BIT 2
   "S_ProgrNo_Bit3_MH06" AT %I71.3 : Bool;   // MH06: preselection program no. MH BIT 3
   "S_ProgrNo_Bit10_MH06" AT %I71.4 : Bool;   // MH06: preselection program no. *10 MH BIT 0
   "S_ProgrNo_Bit20_MH06" AT %I71.5 : Bool;   // MH06: preselection program no. *10 MH BIT 1
   "S_ProgrNo_Bit40_MH06" AT %I71.6 : Bool;   // MH06: preselection program no. *10 MH BIT 2
   "S_ProgrNo_Bit80_MH06" AT %I71.7 : Bool;   // MH06: preselection program no. *10 MH BIT 3
   "S_Manuel_MH06" AT %I72.0 : Bool;   // MH06: operation mode manual
   "S_Automatic_MH06" AT %I72.1 : Bool;   // MH06: operation mode automatic
   "S_Rel_SWU_MH06" AT %I72.2 : Bool;   // MH06: release switch over unit
   "T_CP_forward_MH06" AT %I72.3 : Bool;   // MH06: Button cleaning piston forwards
   "T_CP_back_MH06" AT %I72.4 : Bool;   // MH06: Button cleaning piston back
   "T_Highpressure_MH06" AT %I72.5 : Bool;   // MH06: Button high pressure circulation
   "T_Start_MH06" AT %I72.6 : Bool;   // MH06: Button Start foaming
   "T_Stop_MH06" AT %I72.7 : Bool;   // MH06: Button Stop foaming
   "P_Min_Air_MH06" AT %I73.6 : Bool;   // MH06: Min. Druck Reinigungsluft
   "P_Max_Air_MH06" AT %I73.7 : Bool;   // MH06: Max. Druck Reinigungsluft
   "T_BreakeOpen_MH06" AT %I73.5 : Bool;   // MH06: Button to open the boom brake
   "IPS_MH_MH07" AT %I74.0 : Bool;   // MH06: Inductive proximity switch mixinghead
   "IPS_CP_MH07" AT %I74.1 : Bool;   // MH06: Inductive proximity switch cleaning piston mixinghead
   "ES_OP_Panel_MH07" AT %I74.2 : Bool;   // MH06: Emergency stop operating panel mixinghead
   "K_PreparationFoamingMC07" AT %I74.6 : Bool;   // MH06: preparation foaming from mouldcarrier
   "K_FoamingReleaseMC07" AT %I74.7 : Bool;   // MH06: shot release from mouldcarrier
   "S_ProgNoSelectMH07" AT %IB75 : Byte;   // MH06: preselection program no. MH
   "S_ProgrNo_Bit0_MH07" AT %I75.0 : Bool;   // MH06: preselection program no. MH BIT 0
   "S_ProgrNo_Bit1_MH07" AT %I75.1 : Bool;   // MH06: preselection program no. MH BIT 1
   "S_ProgrNo_Bit2_MH07" AT %I75.2 : Bool;   // MH06: preselection program no. MH BIT 2
   "S_ProgrNo_Bit3_MH07" AT %I75.3 : Bool;   // MH06: preselection program no. MH BIT 3
   "S_ProgrNo_Bit10_MH07" AT %I75.4 : Bool;   // MH06: preselection program no. *10 MH BIT 0
   "S_ProgrNo_Bit20_MH07" AT %I75.5 : Bool;   // MH06: preselection program no. *10 MH BIT 1
   "S_ProgrNo_Bit40_MH07" AT %I75.6 : Bool;   // MH06: preselection program no. *10 MH BIT 2
   "S_ProgrNo_Bit80_MH07" AT %I75.7 : Bool;   // MH06: preselection program no. *10 MH BIT 3
   "S_Manuel_MH07" AT %I76.0 : Bool;   // MH06: operation mode manual
   "S_Automatic_MH07" AT %I76.1 : Bool;   // MH06: operation mode automatic
   "S_Rel_SWU_MH07" AT %I76.2 : Bool;   // MH06: release switch over unit
   "T_CP_forward_MH07" AT %I76.3 : Bool;   // MH06: Button cleaning piston forwards
   "T_CP_back_MH07" AT %I76.4 : Bool;   // MH06: Button cleaning piston back
   "T_Highpressure_MH07" AT %I76.5 : Bool;   // MH06: Button high pressure circulation
   "T_Start_MH07" AT %I76.6 : Bool;   // MH06: Button Start foaming
   "T_Stop_MH07" AT %I76.7 : Bool;   // MH06: Button Stop foaming
   "P_Min_Air_MH07" AT %I77.6 : Bool;   // MH06: Min. Druck Reinigungsluft
   "P_Max_Air_MH07" AT %I77.7 : Bool;   // MH06: Max. Druck Reinigungsluft
   "T_BreakeOpen_MH07" AT %I77.5 : Bool;   // MH06: Button to open the boom brake
   "IPS_MH_MH08" AT %I78.0 : Bool;   // MH06: Inductive proximity switch mixinghead
   "IPS_CP_MH08" AT %I78.1 : Bool;   // MH06: Inductive proximity switch cleaning piston mixinghead
   "ES_OP_Panel_MH08" AT %I78.2 : Bool;   // MH06: Emergency stop operating panel mixinghead
   "K_PreparationFoamingMC08" AT %I78.6 : Bool;   // MH06: preparation foaming from mouldcarrier
   "K_FoamingReleaseMC08" AT %I78.7 : Bool;   // MH06: shot release from mouldcarrier
   "S_ProgNoSelectMH08" AT %IB79 : Byte;   // MH06: preselection program no. MH
   "S_ProgrNo_Bit0_MH08" AT %I79.0 : Bool;   // MH06: preselection program no. MH BIT 0
   "S_ProgrNo_Bit1_MH08" AT %I79.1 : Bool;   // MH06: preselection program no. MH BIT 1
   "S_ProgrNo_Bit2_MH08" AT %I79.2 : Bool;   // MH06: preselection program no. MH BIT 2
   "S_ProgrNo_Bit3_MH08" AT %I79.3 : Bool;   // MH06: preselection program no. MH BIT 3
   "S_ProgrNo_Bit10_MH08" AT %I79.4 : Bool;   // MH06: preselection program no. *10 MH BIT 0
   "S_ProgrNo_Bit20_MH08" AT %I79.5 : Bool;   // MH06: preselection program no. *10 MH BIT 1
   "S_ProgrNo_Bit40_MH08" AT %I79.6 : Bool;   // MH06: preselection program no. *10 MH BIT 2
   "S_ProgrNo_Bit80_MH08" AT %I79.7 : Bool;   // MH06: preselection program no. *10 MH BIT 3
   "S_Manuel_MH08" AT %I80.0 : Bool;   // MH06: operation mode manual
   "S_Automatic_MH08" AT %I80.1 : Bool;   // MH06: operation mode automatic
   "S_Rel_SWU_MH08" AT %I80.2 : Bool;   // MH06: release switch over unit
   "T_CP_forward_MH08" AT %I80.3 : Bool;   // MH06: Button cleaning piston forwards
   "T_CP_back_MH08" AT %I80.4 : Bool;   // MH06: Button cleaning piston back
   "T_Highpressure_MH08" AT %I80.5 : Bool;   // MH06: Button high pressure circulation
   "T_Start_MH08" AT %I80.6 : Bool;   // MH06: Button Start foaming
   "T_Stop_MH08" AT %I80.7 : Bool;   // MH06: Button Stop foaming
   "P_Min_Air_MH08" AT %I81.6 : Bool;   // MH06: Min. Druck Reinigungsluft
   "P_Max_Air_MH08" AT %I81.7 : Bool;   // MH06: Max. Druck Reinigungsluft
   "T_BreakeOpen_MH08" AT %I81.5 : Bool;   // MH06: Button to open the boom brake
   "IPS_MH_MH09" AT %I82.0 : Bool;   // MH06: Inductive proximity switch mixinghead
   "IPS_CP_MH09" AT %I82.1 : Bool;   // MH06: Inductive proximity switch cleaning piston mixinghead
   "ES_OP_Panel_MH09" AT %I82.2 : Bool;   // MH06: Emergency stop operating panel mixinghead
   "K_PreparationFoamingMC09" AT %I82.6 : Bool;   // MH06: preparation foaming from mouldcarrier
   "K_FoamingReleaseMC09" AT %I82.7 : Bool;   // MH06: shot release from mouldcarrier
   "S_ProgNoSelectMH09" AT %IB83 : Byte;   // MH06: preselection program no. MH
   "S_ProgrNo_Bit0_MH09" AT %I83.0 : Bool;   // MH06: preselection program no. MH BIT 0
   "S_ProgrNo_Bit1_MH09" AT %I83.1 : Bool;   // MH06: preselection program no. MH BIT 1
   "S_ProgrNo_Bit2_MH09" AT %I83.2 : Bool;   // MH06: preselection program no. MH BIT 2
   "S_ProgrNo_Bit3_MH09" AT %I83.3 : Bool;   // MH06: preselection program no. MH BIT 3
   "S_ProgrNo_Bit10_MH09" AT %I83.4 : Bool;   // MH06: preselection program no. *10 MH BIT 0
   "S_ProgrNo_Bit20_MH09" AT %I83.5 : Bool;   // MH06: preselection program no. *10 MH BIT 1
   "S_ProgrNo_Bit40_MH09" AT %I83.6 : Bool;   // MH06: preselection program no. *10 MH BIT 2
   "S_ProgrNo_Bit80_MH09" AT %I83.7 : Bool;   // MH06: preselection program no. *10 MH BIT 3
   "S_Manuel_MH09" AT %I84.0 : Bool;   // MH06: operation mode manual
   "S_Automatic_MH09" AT %I84.1 : Bool;   // MH06: operation mode automatic
   "S_Rel_SWU_MH09" AT %I84.2 : Bool;   // MH06: release switch over unit
   "T_CP_forward_MH09" AT %I84.3 : Bool;   // MH06: Button cleaning piston forwards
   "T_CP_back_MH09" AT %I84.4 : Bool;   // MH06: Button cleaning piston back
   "T_Highpressure_MH09" AT %I84.5 : Bool;   // MH06: Button high pressure circulation
   "T_Start_MH09" AT %I84.6 : Bool;   // MH06: Button Start foaming
   "T_Stop_MH09" AT %I84.7 : Bool;   // MH06: Button Stop foaming
   "P_Min_Air_MH09" AT %I85.6 : Bool;   // MH06: Min. Druck Reinigungsluft
   "P_Max_Air_MH09" AT %I85.7 : Bool;   // MH06: Max. Druck Reinigungsluft
   "T_BreakeOpen_MH09" AT %I85.5 : Bool;   // MH06: Button to open the boom brake
   "IPS_MH_MH10" AT %I86.0 : Bool;   // MH06: Inductive proximity switch mixinghead
   "IPS_CP_MH10" AT %I86.1 : Bool;   // MH06: Inductive proximity switch cleaning piston mixinghead
   "ES_OP_Panel_MH10" AT %I86.2 : Bool;   // MH06: Emergency stop operating panel mixinghead
   "K_PreparationFoamingMC10" AT %I86.6 : Bool;   // MH06: preparation foaming from mouldcarrier
   "K_FoamingReleaseMC10" AT %I86.7 : Bool;   // MH06: shot release from mouldcarrier
   "S_ProgNoSelectMH10" AT %IB87 : Byte;   // MH06: preselection program no. MH
   "S_ProgrNo_Bit0_MH10" AT %I87.0 : Bool;   // MH06: preselection program no. MH BIT 0
   "S_ProgrNo_Bit1_MH10" AT %I87.1 : Bool;   // MH06: preselection program no. MH BIT 1
   "S_ProgrNo_Bit2_MH10" AT %I87.2 : Bool;   // MH06: preselection program no. MH BIT 2
   "S_ProgrNo_Bit3_MH10" AT %I87.3 : Bool;   // MH06: preselection program no. MH BIT 3
   "S_ProgrNo_Bit10_MH10" AT %I87.4 : Bool;   // MH06: preselection program no. *10 MH BIT 0
   "S_ProgrNo_Bit20_MH10" AT %I87.5 : Bool;   // MH06: preselection program no. *10 MH BIT 1
   "S_ProgrNo_Bit40_MH10" AT %I87.6 : Bool;   // MH06: preselection program no. *10 MH BIT 2
   "S_ProgrNo_Bit80_MH10" AT %I87.7 : Bool;   // MH06: preselection program no. *10 MH BIT 3
   "S_Manuel_MH10" AT %I88.0 : Bool;   // MH06: operation mode manual
   "S_Automatic_MH10" AT %I88.1 : Bool;   // MH06: operation mode automatic
   "S_Rel_SWU_MH10" AT %I88.2 : Bool;   // MH06: release switch over unit
   "T_CP_forward_MH10" AT %I88.3 : Bool;   // MH06: Button cleaning piston forwards
   "T_CP_back_MH10" AT %I88.4 : Bool;   // MH06: Button cleaning piston back
   "T_Highpressure_MH10" AT %I88.5 : Bool;   // MH06: Button high pressure circulation
   "T_Start_MH10" AT %I88.6 : Bool;   // MH06: Button Start foaming
   "T_Stop_MH10" AT %I88.7 : Bool;   // MH06: Button Stop foaming
   "P_air_2" AT %I19.6 : Bool;   // Pressure air inlet, smooth monitoring
   "P_Max_Air_MH10" AT %I89.7 : Bool;   // MH06: Max. Druck Reinigungsluft
   "T_BreakeOpen_MH10" AT %I89.5 : Bool;   // MH06: Button to open the boom brake
END_VAR
